(* Logix 5000 project; controller PLC_MCC1201_220AP1 vendor 1 type 14 code 164 rev 35.11; software revision 35.00; part 19 of 25 *)
(* tags used below, declared in another part *)
   TMP_xSimulationMode : BOOL;
   AFI : ALIAS FOR B3[7].15;
   AMAX_LEHR_SPD : ALIAS FOR I[81];
   C5 : COUNTER[100];
   C5_ACTIVE_LAMP : ALIAS FOR N54[264].0;
   C5_NTH_IN_LMP : ALIAS FOR N54[264].10;
   C5_NTH_IN_PE : ALIAS FOR N54[264].6;
   C5_NTH_OUT_LMP : ALIAS FOR N54[264].9;
   C5_NTH_OUT_PE : ALIAS FOR N54[264].5;
   C5_STH_IN_LMP : ALIAS FOR N54[264].12;
   C5_STH_IN_PE : ALIAS FOR N54[264].8;
   C5_STH_OUT_LMP : ALIAS FOR N54[264].11;
   C5_STH_OUT_PE : ALIAS FOR N54[264].7;
   CR1_DNET_SS1 : ALIAS FOR N179[18];
   CR1_DNET_SS2 : ALIAS FOR N179[30];
   DRIVE_FAULT_PRESENT : BOOL;
   F96 : REAL[50];
   HMI_Alarm_Presence : BOOL;   // HMI_Alarm_Presence
   HMI_Alarms_0 : BOOL[32];   // HMI Alarms
   HMI_Alarms_1 : BOOL[32];   // HMI Alarms
   HMI_Alarms_2 : BOOL[32];   // HMI Alarms
   HMI_Alarms_3 : BOOL[32];   // HMI Alarms
   HMI_Alarms_4 : BOOL[32];   // HMI Alarms
   HMI_Alarms_5 : BOOL[32];   // HMI Alarms
   HMI_Alarms_6 : BOOL[32];   // HMI Alarms
   HMI_Alarms_7 : BOOL[32];   // HMI Alarms
   HMI_Alarms_8 : BOOL[32];   // HMI Alarms
   HMI_Alarms_9 : BOOL[32];   // HMI Alarms
   HMI_MAN_CMD_WR : UDT_MAN_CMD_WR;
   I : INT[128];
   LEHRSPD_CURRENT : ALIAS FOR N98[5];
   M203DROP : MAC_DROPCONV;
   M205BREAKER : MAC_BREAKER;
   M225 : MAC_EMERGENCYXCUT;
   N11 : DINT[1000];
   N11_HOST : INT[1000];
   N12 : DINT[1000];
   N12_HOST : INT[1000];
   N14 : DINT[1000];
   N14_HOST : INT[1000];
   N179 : DINT[600];
   N500 : DINT[24];
   N501 : DINT[25];
   N502 : DINT[25];
   N504 : DINT[25];
   N505 : DINT[25];
   N507 : DINT[25];
   N53 : DINT[10];
   N53_HOST : INT[10];
   N54 : DINT[501];
   N54_HOST : INT[501];
   O : INT[128];
   ProducedToCullet : UDT_PRODUCED_CULLET;
   ProducedToMCC1300 : UDT_PRODUCED_NEXT;
   R509 : CONTROL[2];
   R509_000_POS : ALIAS FOR R509[0].POS;
   R509_001_POS : ALIAS FOR R509[1].POS;
   S : INT[128];
   Sbr_IN_dDataLength : DINT;
   Status : INT;   // INT tag to retrieve Status value through GSV created during conversion
   T160 : TIMER[100];
   TMP_dIndex : DINT;
   TMP_Index : DINT;
   TMP_xAlwaysOFF : BOOL;
   To_Cullet : DINT[10];
   W_APC_ACTIVE : ALIAS FOR W_B3[0].10;
   W_B3 : DINT[7];
   W_C5 : COUNTER[1];
   W_CB1_AUXILLARY : ALIAS FOR W_I[8].12;
   W_CB1_START : ALIAS FOR W_O[10].1;
   W_CB2_AUXILLARY : ALIAS FOR W_I[8].11;
   W_CB2_START : ALIAS FOR W_O[10].3;
   W_CONV_MSG_N7_0 : MESSAGE;   // IFE1_BTW_CNT
   W_CONV_MSG_N7_120 : MESSAGE;   // OFE1_CONTROL
   W_CONV_MSG_N7_160 : MESSAGE;   // OFE1_BTR_CONTRO
   W_CONV_MSG_N7_200 : MESSAGE;   // OFE2_CONTROL
   W_CONV_MSG_N7_240 : MESSAGE;   // OFE2_BTR_CONTRO
   W_CONV_MSG_N7_280 : MESSAGE;   // OFE3_CONTROL
   W_CONV_MSG_N7_32 : MESSAGE;   // IFE1_BTR
   W_CONV_MSG_N7_320 : MESSAGE;   // OFE3_BTR_CONTRL
   W_CONV_MSG_N7_360 : MESSAGE;   // OFE4_CONTROL
   W_CONV_MSG_N7_400 : MESSAGE;   // OFE4_BTR_CONTRL
   W_CONV_MSG_N7_60 : MESSAGE;   // IFE2_CONTROL
   W_CONV_MSG_N7_92 : MESSAGE;   // IFE2_BTR
   W_CONV_PID_N7_440 : PID;   // Receiving Tank Level Control
   W_CONV_PID_N7_470 : PID;   // Washer Water Pressure Cntrl Valve Position
   W_CONV_PID_N7_500 : PID;   // Dryer Room Airflow (CB2) Fan Actuator Control
   W_CONV_PID_N7_530 : PID;   // Blower CB1 Static Pressure Fan Actuator Control
   W_CONV_PID_N7_560 : PID;   // RO Heating Coil Temp. Control (HC1)
   W_CONV_PID_N7_590 : PID;   // Eclipse Heating Coil Temp. Control
   W_CP1_ENABLE : ALIAS FOR W_B3[0].5;
   W_CP1A_START : ALIAS FOR W_O[10].5;
   W_CP1A_STATUS : ALIAS FOR W_I[8].7;
   W_CP1B_START : ALIAS FOR W_O[10].7;
   W_CP1B_STATUS : ALIAS FOR W_I[8].6;
   W_CP2A_START : ALIAS FOR W_O[10].9;
   W_CP2A_STAT : ALIAS FOR W_I[8].4;
   W_CP2B_START : ALIAS FOR W_O[10].11;
   W_CP2B_STAT : ALIAS FOR W_I[8].3;
   W_DRV_OUTPUT : ALIAS FOR W_N7[380];
   W_DRYER_AIR_FLOW : ALIAS FOR W_N7[108];
   W_EMER_STOP : ALIAS FOR W_I[8].13;
   W_EMER_STOP_LIGHT : ALIAS FOR W_O[10].10;
   W_FLOW_ENABLE : ALIAS FOR W_B3[0].9;
   W_HEATING_AIR_ST : ALIAS FOR W_N7[107];
   W_I : INT[32];
   W_INT_FOR_BCD1 : ALIAS FOR W_N7[911];
   W_LEVEL_SENSOR : ALIAS FOR W_N7[109];
   W_LL_CP1 : ALIAS FOR W_I[8].14;
   W_LL_CP2 : ALIAS FOR W_I[8].15;
   W_LOG_SHUTDOWN : ALIAS FOR W_I[8].0;
   W_N7 : DINT[933];
   W_O : INT[32];
   W_OUT_FROM_PID : ALIAS FOR W_N7[907];
   W_PID_BCD_TCD2 : ALIAS FOR W_N7[913];
   W_PID_TO_OUTPUT : ALIAS FOR W_N7[903];
   W_PS1_SWITCH : ALIAS FOR W_I[8].8;
   W_PWT_HIGH_LIMIT : ALIAS FOR W_I[8].2;
   W_RECIEVING_LEVEL : ALIAS FOR W_I[8].9;
   W_RO_SIG_START : ALIAS FOR W_B3[6].4;
   W_RO_START : ALIAS FOR W_O[10].13;
   W_RUN_WASHER : ALIAS FOR W_B3[0].2;
   W_SHUTDOWN_LATCH : ALIAS FOR W_B3[0].1;
   W_SIG_CP1A_START : ALIAS FOR W_B3[0].6;
   W_SIG_CP1B_START : ALIAS FOR W_B3[0].7;
   W_SIG_CP2A_START : ALIAS FOR W_B3[0].3;
   W_SIG_CP2B_START : ALIAS FOR W_B3[0].4;
   W_T4 : TIMER[101];
   W_TCD1_OUTPUT : ALIAS FOR W_N7[222];
   W_TCD2_OUTPUT : ALIAS FOR W_N7[223];
   W_TT8_INPUT : ALIAS FOR W_N7[912];
   W_TT8_RAW_DATA : ALIAS FOR W_N7[53];
   W_WARNING_LIGHT : ALIAS FOR W_O[10].8;
   Z200 : MAC_Zone_ML;
(* MainProgram, continued *)

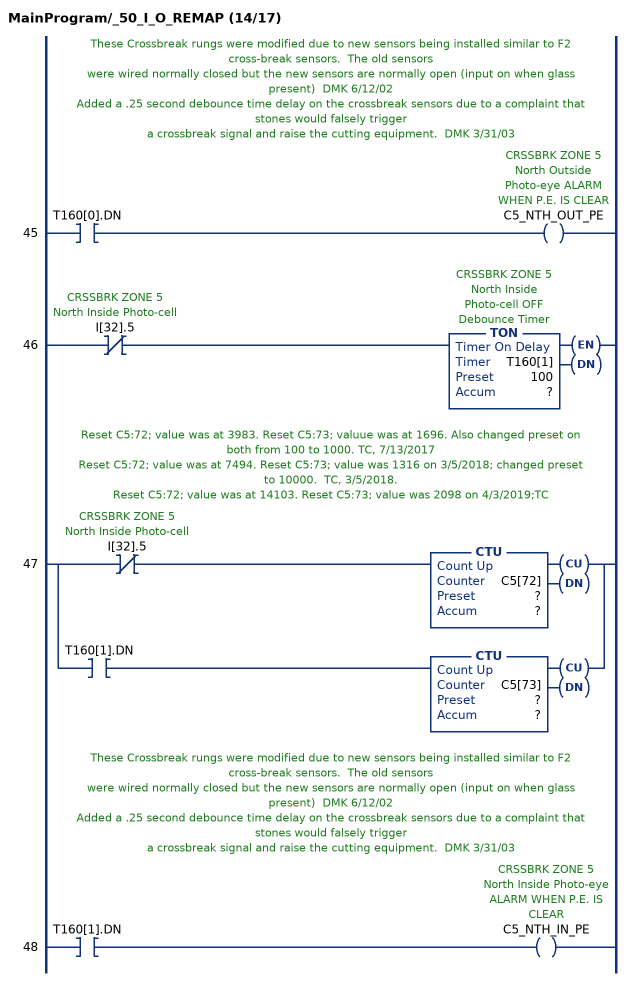
   [picture p306: MainProgram/_50_I_O_REMAP rungs 45-48]
   // These Crossbreak rungs were modified due to new sensors being installed similar to F2 cross-break sensors.  The old sensors
   // were wired normally closed but the new sensors are normally open (input on when glass present)  DMK 6/12/02
   // Added a .25 second debounce time delay on the crossbreak sensors due to a complaint that stones would falsely trigger
   // a crossbreak signal and raise the cutting equipment.  DMK 3/31/03
   45: XIC(T160[0].DN)OTE(C5_NTH_OUT_PE);
   46: XIO(I[32].5)TON(T160[1],?,?);
   // Reset C5:72; value was at 3983. Reset C5:73; valuue was at 1696. Also changed preset on both from 100 to 1000. TC, 7/13/2017
   //                                                                                                                                                       Reset C5:72; value was at 7494. Reset C5:73; value was 1316 on 3/5/2018; changed preset to 10000.  TC, 3/5/2018.
   //                                                                                                                                                                      Reset C5:72; value was at 14103. Reset C5:73; value was 2098 on 4/3/2019;TC
   47: [XIO(I[32].5) CTU(C5[72],?,?) ,XIC(T160[1].DN) CTU(C5[73],?,?) ];
   // These Crossbreak rungs were modified due to new sensors being installed similar to F2 cross-break sensors.  The old sensors
   // were wired normally closed but the new sensors are normally open (input on when glass present)  DMK 6/12/02
   // Added a .25 second debounce time delay on the crossbreak sensors due to a complaint that stones would falsely trigger
   // a crossbreak signal and raise the cutting equipment.  DMK 3/31/03
   48: XIC(T160[1].DN)OTE(C5_NTH_IN_PE);
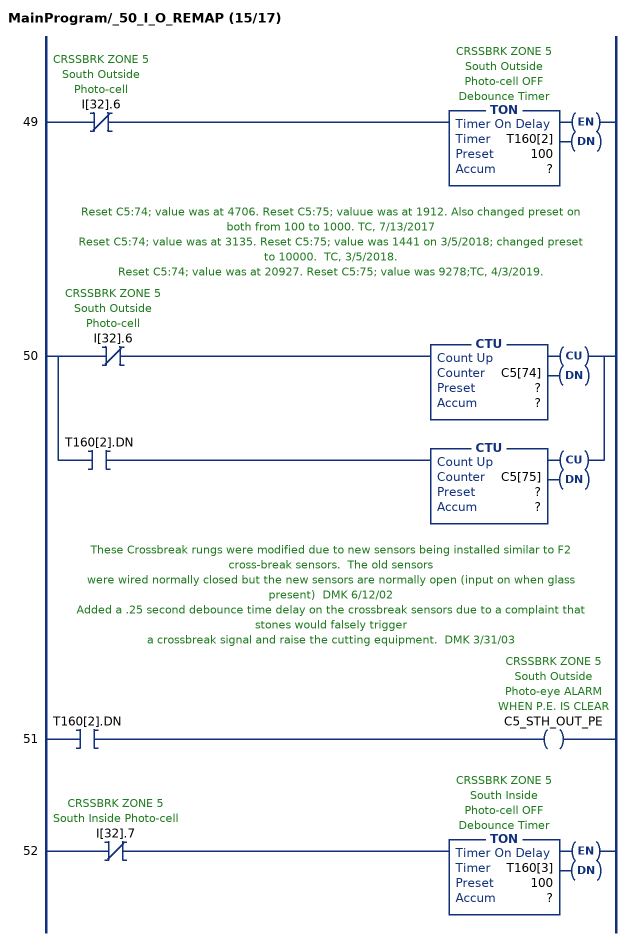
   49: XIO(I[32].6)TON(T160[2],?,?);
   // Reset C5:74; value was at 4706. Reset C5:75; valuue was at 1912. Also changed preset on both from 100 to 1000. TC, 7/13/2017
   //                                                                                                                                                                  Reset C5:74; value was at 3135. Reset C5:75; value was 1441 on 3/5/2018; changed preset to 10000.  TC, 3/5/2018.
   //                                                                                                                                                                                          Reset C5:74; value was at 20927. Reset C5:75; value was 9278;TC, 4/3/2019.
   50: [XIO(I[32].6) CTU(C5[74],?,?) ,XIC(T160[2].DN) CTU(C5[75],?,?) ];
   // These Crossbreak rungs were modified due to new sensors being installed similar to F2 cross-break sensors.  The old sensors
   // were wired normally closed but the new sensors are normally open (input on when glass present)  DMK 6/12/02
   // Added a .25 second debounce time delay on the crossbreak sensors due to a complaint that stones would falsely trigger
   // a crossbreak signal and raise the cutting equipment.  DMK 3/31/03
   51: XIC(T160[2].DN)OTE(C5_STH_OUT_PE);
   52: XIO(I[32].7)TON(T160[3],?,?);
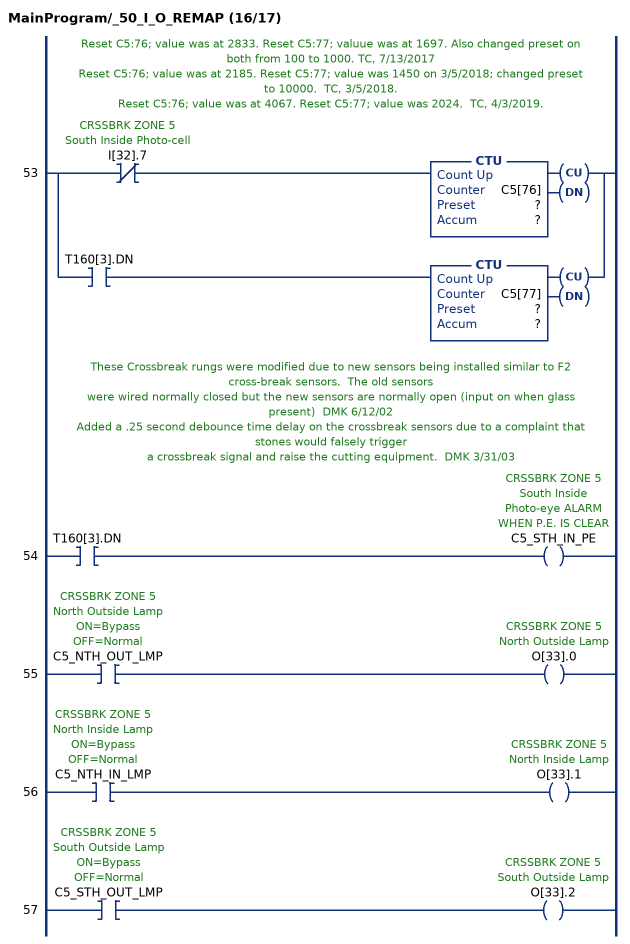
   // Reset C5:76; value was at 2833. Reset C5:77; valuue was at 1697. Also changed preset on both from 100 to 1000. TC, 7/13/2017
   //                                                                                                                                                     Reset C5:76; value was at 2185. Reset C5:77; value was 1450 on 3/5/2018; changed preset to 10000.  TC, 3/5/2018.
   //                                                                                                                                                                               Reset C5:76; value was at 4067. Reset C5:77; value was 2024.  TC, 4/3/2019.
   53: [XIO(I[32].7) CTU(C5[76],?,?) ,XIC(T160[3].DN) CTU(C5[77],?,?) ];
   // These Crossbreak rungs were modified due to new sensors being installed similar to F2 cross-break sensors.  The old sensors
   // were wired normally closed but the new sensors are normally open (input on when glass present)  DMK 6/12/02
   // Added a .25 second debounce time delay on the crossbreak sensors due to a complaint that stones would falsely trigger
   // a crossbreak signal and raise the cutting equipment.  DMK 3/31/03
   54: XIC(T160[3].DN)OTE(C5_STH_IN_PE);
   55: XIC(C5_NTH_OUT_LMP)OTE(O[33].0);
   56: XIC(C5_NTH_IN_LMP)OTE(O[33].1);
   57: XIC(C5_STH_OUT_LMP)OTE(O[33].2);
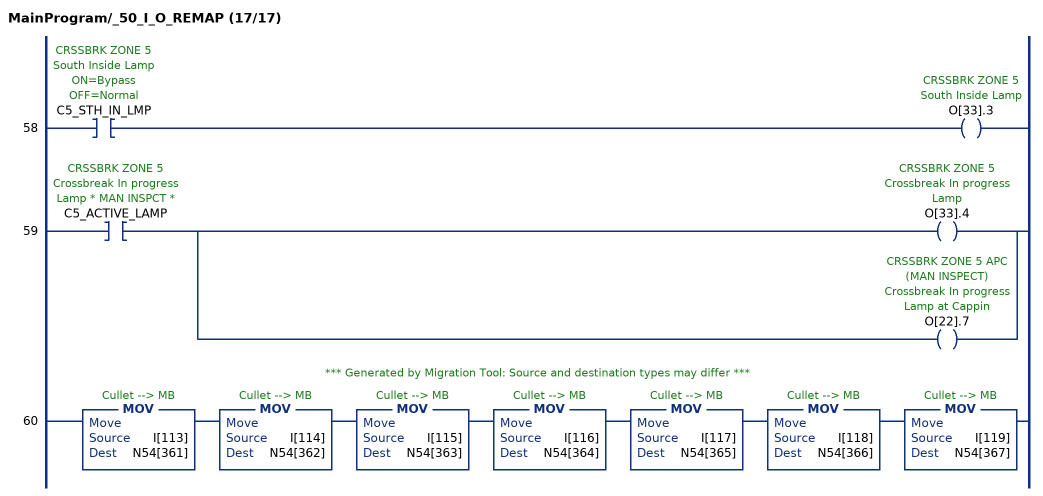
   58: XIC(C5_STH_IN_LMP)OTE(O[33].3);
   59: XIC(C5_ACTIVE_LAMP)[OTE(O[33].4) ,OTE(O[22].7) ];
   // *** Generated by Migration Tool: Source and destination types may differ ***
   60: MOV(I[113],N54[361])MOV(I[114],N54[362])MOV(I[115],N54[363])MOV(I[116],N54[364])MOV(I[117],N54[365])MOV(I[118],N54[366])MOV(I[119],N54[367]);
END_ROUTINE

ROUTINE _51_LADDER   (* ladder *)
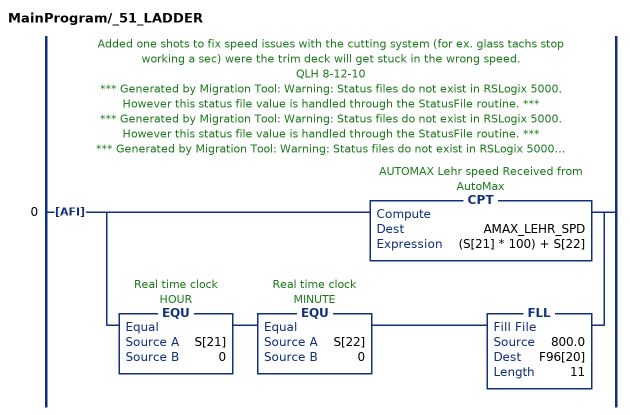
   // Added one shots to fix speed issues with the cutting system (for ex. glass tachs stop working a sec) were the trim deck will get stuck in the wrong speed.
   // QLH 8-12-10
   // *** Generated by Migration Tool: Warning: Status files do not exist in RSLogix 5000. However this status file value is handled through the StatusFile routine. ***
   // *** Generated by Migration Tool: Warning: Status files do not exist in RSLogix 5000. However this status file value is handled through the StatusFile routine. ***
   // *** Generated by Migration Tool: Warning: Status files do not exist in RSLogix 5000. However this status file value is handled through the StatusFile routine. ***
   // *** Generated by Migration Tool: Warning: Status files do not exist in RSLogix 5000. However this status file value is handled through the StatusFile routine. ***
   0: AFI()[CPT(AMAX_LEHR_SPD,(S[21] * 100) + S[22]) ,EQU(S[21],0) EQU(S[22],0) FLL(800.0,F96[20],11) ];
END_ROUTINE

ROUTINE _811_HOST_MOVE   (* structured text *)
   
   //Input
   SBR(Sbr_IN_dDataLength);
   
   FOR TMP_dIndex := 0 TO Sbr_IN_dDataLength - 1 DO
   	N11_HOST[TMP_dIndex] := N11[TMP_dIndex];
   END_FOR;
   
END_ROUTINE

ROUTINE _812_HOST_MOVE   (* structured text *)
   
   //Input
   SBR(Sbr_IN_dDataLength);
   
   FOR TMP_dIndex := 0 TO Sbr_IN_dDataLength - 1 DO
   	N12[TMP_dIndex] := N12_HOST[TMP_dIndex];
   END_FOR;
   
END_ROUTINE

ROUTINE _814_HOST_MOVE   (* structured text *)
   
   
   //Input
   SBR(Sbr_IN_dDataLength);
   
   FOR TMP_dIndex := 0 TO Sbr_IN_dDataLength - 1 DO
   	N14[TMP_dIndex] := N14_HOST[TMP_dIndex];
   END_FOR;
   
END_ROUTINE

ROUTINE _853_HOST_MOVE   (* structured text *)
   
   //Input
   SBR(Sbr_IN_dDataLength);
   
   FOR TMP_dIndex := 0 TO Sbr_IN_dDataLength - 1 DO
   	N53[TMP_dIndex] := N53_HOST[TMP_dIndex];
   END_FOR;
   
END_ROUTINE

ROUTINE _854_HOST_MOVE   (* structured text *)
   
   //Input
   SBR(Sbr_IN_dDataLength);
   
   FOR TMP_dIndex := 0 TO Sbr_IN_dDataLength - 1 DO
   	N54_HOST[TMP_dIndex] := N54[TMP_dIndex];
   END_FOR;
   
END_ROUTINE

ROUTINE _880_HMI_Mapping   (* structured text *)
   
   // Alarm maps for HMI
   TMP_Index:= 0;
   FOR TMP_Index := 0 TO 15 DO
   	//HMI_Alarms_0[TMP_Index]:= N11[62].[TMP_Index];
   	//HMI_Alarms_1[TMP_Index]:= N11[64].[TMP_Index];
   	HMI_Alarms_0[TMP_Index]:= 0;
   	HMI_Alarms_1[TMP_Index]:= 0;
   	HMI_Alarms_2[TMP_Index]:= 0;
   	HMI_Alarms_3[TMP_Index]:= 0;
   	HMI_Alarms_4[TMP_Index]:= 0;
   	HMI_Alarms_5[TMP_Index]:= 0;
   	HMI_Alarms_6[TMP_Index]:= 0;
   	HMI_Alarms_7[TMP_Index]:= 0;
   	HMI_Alarms_8[TMP_Index]:= 0;
   	HMI_Alarms_9[TMP_Index]:= 0;
   	//HMI_Alarms_2[TMP_Index]:= NOT N11[22].[TMP_Index];
   	//HMI_Alarms_3[TMP_Index]:= NOT N11[23].[TMP_Index];
   END_FOR;
   FOR TMP_Index := 16 TO 31 DO
   	HMI_Alarms_0[TMP_Index]:= 0;
   	HMI_Alarms_1[TMP_Index]:= 0;
   	HMI_Alarms_2[TMP_Index]:= 0;
   	HMI_Alarms_3[TMP_Index]:= 0;
   	HMI_Alarms_4[TMP_Index]:= 0;
   	HMI_Alarms_5[TMP_Index]:= 0;
   	HMI_Alarms_6[TMP_Index]:= 0;
   	HMI_Alarms_7[TMP_Index]:= 0;
   	HMI_Alarms_8[TMP_Index]:= 0;
   	HMI_Alarms_9[TMP_Index]:= 0;
   END_FOR;
   
   (*
   HMI_Alarms_0[0] := NOT N11[20].0;
   HMI_Alarms_0[1] := NOT N11[20].1;
   HMI_Alarms_0[2] := NOT N11[20].2;
   HMI_Alarms_0[3] := NOT N11[20].3;
   HMI_Alarms_0[4] := 0;
   HMI_Alarms_0[5] := NOT N11[20].5;
   HMI_Alarms_0[6] := NOT N11[20].6;
   HMI_Alarms_0[7] := NOT N11[20].7;
   HMI_Alarms_0[8] := N11[20].8;
   HMI_Alarms_0[9] := N11[20].9;
   HMI_Alarms_0[10] := NOT N11[20].10;
   HMI_Alarms_0[11] := NOT N11[20].11;
   HMI_Alarms_0[12] := NOT N11[20].12;
   HMI_Alarms_0[13] := NOT N11[20].13;
   HMI_Alarms_0[14] := N11[20].14;
   HMI_Alarms_0[15] := 0;
   
   HMI_Alarms_2[0] := NOT N11[22].0;
   HMI_Alarms_2[1] := NOT N11[22].1;
   HMI_Alarms_2[2] := NOT N11[22].2;
   HMI_Alarms_2[3] := NOT N11[22].3;
   HMI_Alarms_2[4] := NOT N11[22].4;
   HMI_Alarms_2[5] := NOT N11[22].5;
   HMI_Alarms_2[6] := NOT N11[22].6;
   HMI_Alarms_2[7] := NOT N11[22].7;
   HMI_Alarms_2[8] := NOT N11[22].8;
   HMI_Alarms_2[9] := NOT N11[22].9;
   HMI_Alarms_2[10] := NOT N11[22].10;
   HMI_Alarms_2[11] := NOT N11[22].11;
   HMI_Alarms_2[12] := NOT N11[22].12;
   HMI_Alarms_2[13] := NOT N11[22].13;
   HMI_Alarms_2[14] := 0;
   HMI_Alarms_2[15] := 0;
   
   HMI_Alarms_3[0] := NOT N11[23].0;
   HMI_Alarms_3[1] := NOT N11[23].1;
   HMI_Alarms_3[2] := NOT N11[23].2;
   HMI_Alarms_3[3] := NOT N11[23].3;
   HMI_Alarms_3[4] := NOT N11[23].4;
   HMI_Alarms_3[5] := NOT N11[23].5;
   HMI_Alarms_3[6] := NOT N11[23].6;
   HMI_Alarms_3[7] := NOT N11[23].7;
   HMI_Alarms_3[8] := NOT N11[23].8;
   HMI_Alarms_3[9] := NOT N11[23].9;
   HMI_Alarms_3[10] := NOT N11[23].10;
   HMI_Alarms_3[11] := NOT N11[23].11;
   HMI_Alarms_3[12] := NOT N11[23].12;
   HMI_Alarms_3[13] := NOT N11[23].13;
   HMI_Alarms_3[14] := 0;
   HMI_Alarms_3[15] := 0;
   
   HMI_Alarms_9[0] := M316M1_IN.Faulted;
   HMI_Alarms_9[1] := M317M1_IN.Faulted;
   HMI_Alarms_9[2] := M317M2_IN.Faulted;
   HMI_Alarms_9[3] := M317M3_IN.Faulted;
   HMI_Alarms_9[4] := M317M4_IN.Faulted;
   HMI_Alarms_9[5] := M317M5_IN.Faulted;
   HMI_Alarms_9[6] := M317M6_IN.Faulted;
   HMI_Alarms_9[7] := M318M1_IN.Faulted;
   HMI_Alarms_9[8] := M318AM1_IN.Faulted;
   HMI_Alarms_9[9] := M318BM1_IN.Faulted;
   HMI_Alarms_9[10] := M318BM2_IN.Faulted;
   HMI_Alarms_9[11] := M318BM3_IN.Faulted;
   HMI_Alarms_9[12] := M318BM4_IN.Faulted;
   HMI_Alarms_9[13] := M391M1_IN.Faulted;
   *)
   
   // Alarm presence for HMI
   HMI_Alarm_Presence := 0;
   TMP_Index:= 0;
   FOR TMP_Index := 0 TO 31 DO
   	IF HMI_Alarms_0[TMP_Index] OR HMI_Alarms_1[TMP_Index] OR HMI_Alarms_2[TMP_Index] OR HMI_Alarms_3[TMP_Index] OR HMI_Alarms_4[TMP_Index] OR HMI_Alarms_5[TMP_Index] THEN
   		HMI_Alarm_Presence := 1;
   	END_IF;
   	IF HMI_Alarms_6[TMP_Index] OR HMI_Alarms_7[TMP_Index] OR HMI_Alarms_8[TMP_Index] OR HMI_Alarms_9[TMP_Index] THEN
   		HMI_Alarm_Presence := 1;
   	END_IF;
   END_FOR;
   
   //// Logic to make horn sound for drives fault
   //DRIVE_FAULT_PRESENT := 0;
   //FOR TMP_Index := 0 TO 8 BY 1 DO
   //	IF N11[62].[TMP_Index] THEN
   //		DRIVE_FAULT_PRESENT := 1;
   //	END_IF;
   //END_FOR;
   
   (*
   // Photocell maps for HMI
   HMI_ProxySwitch[0] := I[2].0;
   HMI_ProxySwitch[1] := I[2].1;
   HMI_ProxySwitch[2] := I[2].2;
   HMI_ProxySwitch[3] := I[2].3;
   HMI_ProxySwitch[4] := I[2].4;
   HMI_ProxySwitch[5] := I[2].5;
   HMI_ProxySwitch[6] := I[2].6;
   HMI_ProxySwitch[7] := I[2].7;
   HMI_ProxySwitch[8] := I[2].8;
   HMI_ProxySwitch[9] := I[2].9;
   HMI_ProxySwitch[10] := I[2].10;
   HMI_ProxySwitch[11] := I[2].11;
   HMI_ProxySwitch[12] := I[2].12;
   HMI_ProxySwitch[13] := I[2].13;
   HMI_ProxySwitch[14] := I[2].14;
   HMI_ProxySwitch[15] := I[2].15;
   
   // Photocell maps for HMI
   HMI_Photocells[0] := I[3].0;
   HMI_Photocells[1] := I[3].1;
   HMI_Photocells[2] := I[3].2;
   HMI_Photocells[3] := I[3].3;
   HMI_Photocells[4] := I[3].4;
   HMI_Photocells[5] := I[3].5;
   HMI_Photocells[6] := I[3].6;
   HMI_Photocells[7] := I[3].7;
   HMI_Photocells[8] := I[3].8;
   HMI_Photocells[9] := I[3].9;
   HMI_Photocells[10] := I[3].10;
   HMI_Photocells[11] := I[3].11;
   HMI_Photocells[12] := I[3].12;
   HMI_Photocells[13] := I[3].13;
   HMI_Photocells[14] := I[3].14;
   HMI_Photocells[15] := I[3].15;
   
   HMI_Photocells[16] := I[5].8;
   HMI_Photocells[17] := I[5].9;
   
   //All commands
   I[21].15 := HMI_MAN_CMD_WR.CONV_Manual_ALL;
   I[23].15 := HMI_MAN_CMD_WR.CONV_Man_ALL_FWD;
   I[25].15 := HMI_MAN_CMD_WR.CONV_Man_ALL_REV;
   
   //M316M1 Roll Conveyor M4CM01
   I[20].0 := HMI_MAN_CMD_WR.M316M1_Manual;
   I[22].0 := HMI_MAN_CMD_WR.M316M1_ManFWD;
   I[24].0 := HMI_MAN_CMD_WR.M316M1_ManREV;
   
   //M317M1 Roll Conveyor Zone 1 M4CM02
   I[20].1 := HMI_MAN_CMD_WR.M317M1_Manual;
   I[22].1 := HMI_MAN_CMD_WR.M317M1_ManFWD;
   I[24].1 := HMI_MAN_CMD_WR.M317M1_ManREV;
   
   //M317M2 Lifting Zone 1 M4CM03
   I[20].2 := HMI_MAN_CMD_WR.M317M2_Manual;
   I[22].2 := HMI_MAN_CMD_WR.M317M2_ManFWD;
   I[24].2 := HMI_MAN_CMD_WR.M317M2_ManREV;
   
   //M317M3 Lifting Zone 2 M4CM04
   I[20].3 := HMI_MAN_CMD_WR.M317M3_Manual;
   I[22].3 := HMI_MAN_CMD_WR.M317M3_ManFWD;
   I[24].3 := HMI_MAN_CMD_WR.M317M3_ManREV;
   
   //M317M4 Roll Conveyor Zone 2 M4CM05
   I[20].4 := HMI_MAN_CMD_WR.M317M4_Manual;
   I[22].4 := HMI_MAN_CMD_WR.M317M4_ManFWD;
   I[24].4 := HMI_MAN_CMD_WR.M317M4_ManREV;
   
   //M317M5 Wheel Conveyor Zone 1 M4CM06
   I[20].5 := HMI_MAN_CMD_WR.M317M5_Manual;
   I[22].5 := HMI_MAN_CMD_WR.M317M5_ManFWD;
   I[24].5 := HMI_MAN_CMD_WR.M317M5_ManREV;
   
   //M317M6 Wheel Conveyor Zone 2 M4CM07
   I[20].6 := HMI_MAN_CMD_WR.M317M6_Manual;
   I[22].6 := HMI_MAN_CMD_WR.M317M6_ManFWD;
   I[24].6 := HMI_MAN_CMD_WR.M317M6_ManREV;
   
   //M318M1 Roll Conveyor M4CM08
   I[20].7 := HMI_MAN_CMD_WR.M318M1_Manual;
   I[22].7 := HMI_MAN_CMD_WR.M318M1_ManFWD;
   I[24].7 := HMI_MAN_CMD_WR.M318M1_ManREV;
   
   //M318AM1 Roll Conveyor M4CM09
   I[20].8 := HMI_MAN_CMD_WR.M318AM1_Manual;
   I[22].8 := HMI_MAN_CMD_WR.M318AM1_ManFWD;
   I[24].8 := HMI_MAN_CMD_WR.M318AM1_ManREV;
   
   //M318BM1 Roll Conveyor Zone 1 M4CM10
   I[20].9 := HMI_MAN_CMD_WR.M318BM1_Manual;
   I[22].9 := HMI_MAN_CMD_WR.M318BM1_ManFWD;
   I[24].9 := HMI_MAN_CMD_WR.M318BM1_ManREV;
   
   //M318BM2 Lifting Zone 1 M4CM11
   I[20].10 := HMI_MAN_CMD_WR.M318BM2_Manual;
   I[22].10 := HMI_MAN_CMD_WR.M318BM2_ManFWD;
   I[24].10 := HMI_MAN_CMD_WR.M318BM2_ManREV;
   
   //M318BM3 Lifting Zone 2 M4CM12
   I[20].11 := HMI_MAN_CMD_WR.M318BM3_Manual;
   I[22].11 := HMI_MAN_CMD_WR.M318BM3_ManFWD;
   I[24].11 := HMI_MAN_CMD_WR.M318BM3_ManREV;
   
   //M318BM4 Roll Conveyor Zone 2 M4CM13
   I[20].12 := HMI_MAN_CMD_WR.M318BM4_Manual;
   I[22].12 := HMI_MAN_CMD_WR.M318BM4_ManFWD;
   I[24].12 := HMI_MAN_CMD_WR.M318BM4_ManREV;
   
   //M391M1 Wheel Conveyor (Sample Table) M4CM14
   I[20].13 := HMI_MAN_CMD_WR.M391M1_Manual;
   I[22].13 := HMI_MAN_CMD_WR.M391M1_ManFWD;
   I[24].13 := HMI_MAN_CMD_WR.M391M1_ManREV;
   I[22].14 := HMI_MAN_CMD_WR.M391_ManRAISE;
   I[24].14 := HMI_MAN_CMD_WR.M391_ManLOWER;
   *)
   
END_ROUTINE

ROUTINE _990_Output_Mapping   (* structured text *)
   
   //OUTPUT
   
   //MCC1201
   A152AP1:14:O.Pt00.Data := Z200.OUTPUT_xMainEmergencyLamp;
   A152AP1:14:O.Pt01.Data := Z200.OUTPUT_xUPSEmergencyLamp;
   A152AP1:14:O.Pt02.Data := Z200.OUTPUT_xMCCSafetyLamp;
   
   //Alarms signalling
   A152AP1:15:O.Pt03.Data := Z200.OUTPUT_xUPSEmergencyLamp;
   A152AP1:15:O.Pt06.Data := Z200.OUTPUT_xAcousticAlarm;
   A152AP1:15:O.Pt07.Data := Z200.OUTPUT_xUPSEmergencyLamp;
   A152AP1:15:O.Pt11.Data := Z200.OUTPUT_xMainEmergencyLamp;
   A152AP1:15:O.Pt12.Data := Z200.OUTPUT_xMainEmergencyLamp;
   A152AP1:16:O.Pt01.Data := Z200.OUTPUT_xUPSEmergencyLamp;
   A152AP1:16:O.Pt11.Data := Z200.OUTPUT_xUPSEmergencyLamp;
   
   //M203DROP
   A152AP1:15:O.Pt00.Data := M203DROP.OUTPUT_xRollerLifting;
   A152AP1:15:O.Pt01.Data := M203DROP.OUTPUT_xDescentDrop;
   A152AP1:15:O.Pt02.Data := M203DROP.OUTPUT_xRiseDrop;
   A152AP1:15:O.Pt04.Data := M203DROP.OUTPUT_xHLDoorOpenOpSide;
   A152AP1:15:O.Pt05.Data := M203DROP.OUTPUT_xHLUpDownPushbutton;
   A152AP1:15:O.Pt08.Data := M203DROP.OUTPUT_xHLDoorOpenFarSide;
   A152AP1:15:O.Pt09.Data := M203DROP.OUTPUT_xHLUpDownPushbutton;
   
   //M225 EMERGENCY XCUT
   A152AP1:16:O.Pt00.Data := M225.OUTPUT_xUnlockDoorOpSide;
   A152AP1:16:O.Pt02.Data := M225.OUTPUT_xAreaAccessRequestFarSide;
   A152AP1:16:O.Pt05.Data := M225.OUTPUT_xUnlockDoorFarSide;
   A152AP1:16:O.Pt06.Data := M225.OUTPUT_xMachineReady;
   A152AP1:16:O.Pt07.Data := M225.OUTPUT_xMachineToMaintenance;
   A152AP1:16:O.Pt08.Data := M225.OUTPUT_xMachineOutOfOrder;
   A152AP1:18:O.Pt00.Data := M225.OUTPUT_xCuttingHeadDescent;
   A152AP1:18:O.Pt01.Data := M225.OUTPUT_xLubrication;
   A152AP1:18:O.Pt02.Data := M225.OUTPUT_xAirActivation;
   
   //CS4225 EMERGENCY XCUT CONSOLLE
   A152AP1:16:O.Pt12.Data := M225.OUTPUT_xAreaAccessRequestOpSide;
   A152AP1:16:O.Pt13.Data := M225.OUTPUT_xAutomatic;
   A152AP1:16:O.Pt14.Data := M225.OUTPUT_xStartCut;
   A152AP1:16:O.Pt15.Data := M225.OUTPUT_xStopCut;
   
   //M205BREAKER
   A152AP1:13:O.Pt00.Data := M205BREAKER.OUTPUT_xBreakerRun;
   
   //M225
   A152AP1:13:O.Pt01.Data := M225.OUTPUT_xCarriageOverstroke;
   
   
   // MAPPING PREVIOUS PROGRAM OUTPUTS
   
   //HORN / CHILLED WATER / APC / SUBSURFACE / ISRA 5D
   A152AP1:14:O.Pt03.Data := I[20].3; //PLC ALARM HORN RELAY
   A152AP1:14:O.Pt04.Data := I[20].4; //North Chilled Water Blower Start VFD
   A152AP1:14:O.Pt05.Data := I[20].5; //North Chilled Water Blower Start LT I02104 PB
   A152AP1:14:O.Pt06.Data := I[20].6; //North Chilled Water VFD Stop
   A152AP1:14:O.Pt07.Data := I[20].0; //South Chilled Water Blower Start VFD
   A152AP1:14:O.Pt08.Data := I[20].1; //South Chilled Water Blower Start LT I02112 PB
   A152AP1:14:O.Pt09.Data := I[20].2; //South Chilled Water VFD Stop
   A152AP1:14:O.Pt10.Data := I[20].8; //LUCOR MACHINE OPERATE (APC CONTACTORS?)
   A152AP1:14:O.Pt11.Data := I[20].11; //SUB-SURFACE Cutters Raise for Crossbreak Relay
   A152AP1:14:O.Pt12.Data := I[20].12; //ISRA 5D System Cut Signal
   A152AP1:14:O.Pt13.Data := I[20].13; //ISRA 5D System QC Request Signal
   
   // CROSSBREAK ZONE 1
   CB_1CS:1:O.0 := O[25].0; //CRSSBRK ZONE 1 North Outside Lamp
   CB_1CS:1:O.1 := O[25].1; //CRSSBRK ZONE 1 North Inside Lamp
   CB_1CS:1:O.2 := O[25].2; //CRSSBRK ZONE 1 South Outside Lamp
   CB_1CS:1:O.3 := O[25].3; //CRSSBRK ZONE 1 South Inside Lamp
   CB_1CS:1:O.4 := O[25].4; //CRSSBRK ZONE 1 Crossbreak In progress Lamp
   CB_1CS:1:O.5 := O[25].5; //M37B Conv Forward Pilot Light
   CB_1CS:1:O.6 := O[25].6; //M37B Conv Reverse Pilot Light
   CB_1CS:1:O.7 := O[25].7; //M47B Conv Forward Pilot Light
   CB_1CS:1:O.8 := O[25].8; //M47B Conv Reverse Pilot Light
   CB_1CS:1:O.9 := O[25].9; //spare
   CB_1CS:1:O.10 := O[25].10; //spare
   CB_1CS:1:O.11 := O[25].11; //spare
   CB_1CS:1:O.12 := O[25].12; //spare
   CB_1CS:1:O.13 := O[25].13; //spare
   CB_1CS:1:O.14 := O[25].14; //spare
   CB_1CS:1:O.15 := O[25].15; //spare
   
   // CROSSBREAK ZONE 2
   CB_2CS:1:O.0 := O[27].0; //CRSSBRK ZONE 2 North Outside Lamp
   CB_2CS:1:O.1 := O[27].1; //CRSSBRK ZONE 2 North Inside Lamp
   CB_2CS:1:O.2 := O[27].2; //CRSSBRK ZONE 2 South Outside Lamp (Bad Output)
   CB_2CS:1:O.3 := O[27].3; //CRSSBRK ZONE 2 South Inside Lamp
   CB_2CS:1:O.4 := O[27].4; //CRSSBRK ZONE 2 Crossbreak In progress Lamp
   CB_2CS:1:O.5 := O[27].5; //CRSSBRK ZONE 1 Crossbreak horn Located on wall At lehr Exit
   CB_2CS:1:O.6 := O[27].6; //CRSSBRK ZONE 1 Alarm rotating Beacon Located on lehr Exit
   CB_2CS:1:O.7 := O[27].7; //Crusher #1 Is Lowered (This Output is Read by HE for Pan-alarm Display)
   CB_2CS:1:O.8 := O[27].8; //CRSSBRK ZONE 2 South Outside Lamp (New Output)
   CB_2CS:1:O.9 := O[27].9; //spare
   CB_2CS:1:O.10 := O[27].10; //spare
   CB_2CS:1:O.11 := O[27].11; //spare
   CB_2CS:1:O.12 := O[27].12; //spare
   CB_2CS:1:O.13 := O[27].13; //spare
   CB_2CS:1:O.14 := O[27].14; //spare
   CB_2CS:1:O.15 := O[27].15; //spare
   
   // CROSSBREAK ZONE 3
   CB_3CS:1:O.0 := O[29].0; //CRSSBRK ZONE 3 North Outside Lamp
   CB_3CS:1:O.1 := O[29].1; //CRSSBRK ZONE 3 North Inside Lamp
   CB_3CS:1:O.2 := O[29].2; //CRSSBRK ZONE 3 South Outside Lamp (Bad Output)
   CB_3CS:1:O.3 := O[29].3; //CRSSBRK ZONE 3 South Inside Lamp
   CB_3CS:1:O.4 := O[29].4; //CRSSBRK ZONE 3 Crossbreak In progress Lamp
   CB_3CS:1:O.5 := O[29].5; //spare
   CB_3CS:1:O.6 := O[29].6; //spare
   CB_3CS:1:O.7 := O[29].7; //spare
   CB_3CS:1:O.8 := O[29].8; //spare
   CB_3CS:1:O.9 := O[29].9; //spare
   CB_3CS:1:O.10 := O[29].10; //spare
   CB_3CS:1:O.11 := O[29].11; //spare
   CB_3CS:1:O.12 := O[29].12; //spare
   CB_3CS:1:O.13 := O[29].13; //spare
   CB_3CS:1:O.14 := O[29].14; //spare
   CB_3CS:1:O.15 := O[29].15; //spare
   
   // CROSSBREAK ZONE 4 (IMAGE AUTO)
   CB_4CS:1:O.0 := O[31].0; //CRSSBRK ZONE 4 North Outside Lamp
   CB_4CS:1:O.1 := O[31].1; //CRSSBRK ZONE 4 North Inside Lamp
   CB_4CS:1:O.2 := O[31].2; //CRSSBRK ZONE 4 South Outside Lamp (Bad Output)
   CB_4CS:1:O.3 := O[31].3; //CRSSBRK ZONE 4 South Inside Lamp
   CB_4CS:1:O.4 := O[31].4; //CRSSBRK ZONE 4 Crossbreak In progress Lamp
   CB_4CS:1:O.5 := O[31].5; //spare
   CB_4CS:1:O.6 := O[31].6; //IMAGE AUTO Retro cover Manual  mode Lamp
   CB_4CS:1:O.7 := O[31].7; //IMAGE AUTO Retro cover Closed Alarm Horn
   CB_4CS:1:O.8 := O[31].8; //IMAGE AUTO Retro cover Alarm Beacon
   CB_4CS:1:O.9 := O[31].9; //IMAGE AUTO Open Graticule Solenoid (Raise)
   CB_4CS:1:O.10 := O[31].10; //IMAGE AUTO Retro Cover Open solenoid Valve
   CB_4CS:1:O.11 := O[31].11; //spare
   CB_4CS:1:O.12 := O[31].12; //spare
   CB_4CS:1:O.13 := O[31].13; //spare
   CB_4CS:1:O.14 := O[31].14; //spare
   CB_4CS:1:O.15 := O[31].15; //spare
   
   // CROSSBREAK ZONE 5 (APC)
   CB_5CS:1:O.0 := O[33].0; //CRSSBRK ZONE 5 North Outside Lamp
   CB_5CS:1:O.1 := O[33].1; //CRSSBRK ZONE 5 North Inside Lamp
   CB_5CS:1:O.2 := O[33].2; //CRSSBRK ZONE 5 South Outside Lamp (Bad Output)
   CB_5CS:1:O.3 := O[33].3; //CRSSBRK ZONE 5 South Inside Lamp
   CB_5CS:1:O.4 := O[33].4; //CRSSBRK ZONE 5 Crossbreak In progress Lamp
   CB_5CS:1:O.5 := O[33].5; //APC Enable Relay
   CB_5CS:1:O.6 := O[33].6; //APC Cut Off relay New Apc Sprayer
   CB_5CS:1:O.7 := O[33].7; //APC #2 Blow off Excess APC During Crossbreak
   CB_5CS:1:O.8 := O[33].8; //APC #2 Lower Roll (On Glass)
   CB_5CS:1:O.9 := O[33].9; //APC #1 Blow off Excess APC During Crossbreak changed 22Mar2019TC
   CB_5CS:1:O.10 := O[33].10; //APC #1 Lower Roll (On Glass) new22MarTC
   CB_5CS:1:O.11 := O[33].11; //APC APC Roll SS1 changed 22Mar2019TC
   CB_5CS:1:O.12 := O[33].12; //spare
   CB_5CS:1:O.13 := O[33].13; //spare
   CB_5CS:1:O.14 := O[33].14; //spare
   CB_5CS:1:O.15 := O[33].15; //spare
   
   // MANUAL INSPECTION
   MI_6CS:1:O.0 := O[35].0; //MANUAL INSPCTN North Outside Reject Flaw Red Lamp
   MI_6CS:1:O.1 := O[35].1; //MANUAL INSPCTN North Outside Q.A. Flaw Yellow Lamp
   MI_6CS:1:O.2 := O[35].2; //MANUAL INSPCTN North Inside Reject Flaw Red Lamp
   MI_6CS:1:O.3 := O[35].3; //MANUAL INSPCTN North Inside Q.A. Flaw Yellow Lamp
   MI_6CS:1:O.4 := O[35].4; //MANUAL INSPCTN * Center Reject Flaw Red Lamp
   MI_6CS:1:O.5 := O[35].5; //MANUAL INSPCTN * Center Q.A. Flaw Yellow Lamp
   MI_6CS:1:O.6 := O[35].6; //MANUAL INSPCTN South Inside Reject Flaw Red Lamp
   MI_6CS:1:O.7 := O[35].7; //MANUAL INSPCTN South Inside Q.A. Flaw Yellow Lamp
   MI_6CS:1:O.8 := O[35].8; //MANUAL INSPCTN South Outside Reject Flaw Red Lamp
   MI_6CS:1:O.9 := O[35].9; //MANUAL INSPCTN South Outside Q.A. Flaw Yellow Lamp
   MI_6CS:1:O.10 := O[35].10; //MANUAL INSPCTN Cross-break Signal to STP
   MI_6CS:1:O.11 := O[35].11; //spare
   MI_6CS:1:O.12 := O[35].12; //spare
   MI_6CS:1:O.13 := O[35].13; //MANUAL INSPCTN * * Function Lamp Clear
   MI_6CS:1:O.14 := O[35].14; //MANUAL INSPCTN * * Function Lamp Blue
   MI_6CS:1:O.15 := O[35].15; //MANUAL INSPCTN Quality Defect Inhibit Function Lamp Red
   
   //Cabinet
   A152AP1:15:O.Pt15.Data := TMP_xSimulationMode; //PLC ANOMALY
   A152AP1:17:O.Pt00.Data := O[35].15; //MANUAL INSPECTION
   
   //VMCC W1 (WASHER)
   
   
   
   //PANEL W2 (WASHER)
   PANEL_W2:3:O.0 := O[59].0; //PANEL W2 BRUSH #1 Manual mode Lamp
   PANEL_W2:3:O.1 := O[59].1; //SPARE
   PANEL_W2:3:O.2 := O[59].2; //PANEL W2 SPONGE UNIT Manual mode Lamp
   PANEL_W2:3:O.3 := O[59].3; //PANEL W2 AIR KNIVES Manual mode Lamp
   PANEL_W2:3:O.4 := O[59].4; //PANEL W2 WATER SPRAYERS Manual mode Lamp
   PANEL_W2:3:O.5 := O[59].5; //SPARE
   PANEL_W2:3:O.6 := O[59].6; //PANEL W2 AIR KNIFE SS LIGHT ON PANEL #W2
   PANEL_W2:3:O.7 := O[59].7; //PANEL W2 AIR KNIFE RELAY AKBR-ON
   PANEL_W2:3:O.8 := O[59].8; //SPARE
   PANEL_W2:3:O.9 := O[59].9; //SPARE
   PANEL_W2:3:O.10 := O[59].10; //SPARE
   PANEL_W2:3:O.11 := O[59].11; //SPARE
   PANEL_W2:3:O.12 := O[59].12; //SPARE
   PANEL_W2:3:O.13 := O[59].13; //SPARE
   PANEL_W2:3:O.14 := O[59].14; //SPARE
   PANEL_W2:3:O.15 := O[59].15; //SPARE
   
   //PANEL W3 (WASHER)
   PANEL_W3:3:O.0 := O[63].0; //PANEL W3 BRUSH #1 Manual mode Lamp
   PANEL_W3:3:O.1 := O[63].1; //SPARE
   PANEL_W3:3:O.2 := O[63].2; //PANEL W3 SPONGE UNIT Manual mode Lamp
   PANEL_W3:3:O.3 := O[63].3; //PANEL W3 AIR KNIVES Manual mode Lamp
   PANEL_W3:3:O.4 := O[63].4; //PANEL W3 WATER SPRAYERS Manual mode Lamp
   PANEL_W3:3:O.5 := O[63].5; //SPARE
   PANEL_W3:3:O.6 := O[63].6; //PANEL W3 AIR KNIFE SS LIGHT ON PANEL #W3
   PANEL_W3:3:O.7 := O[63].7; //SPARE
   PANEL_W3:3:O.8 := O[63].8; //SPARE
   PANEL_W3:3:O.9 := O[63].9; //SPARE
   PANEL_W3:3:O.10 := O[63].10; //SPARE
   PANEL_W3:3:O.11 := O[63].11; //SPARE
   PANEL_W3:3:O.12 := O[63].12; //SPARE
   PANEL_W3:3:O.13 := O[63].13; //SPARE
   PANEL_W3:3:O.14 := O[63].14; //SPARE
   PANEL_W3:3:O.15 := O[63].15; //SPARE
   
   
   //PRODUCED
   
   To_Cullet[0] := O[112];
   To_Cullet[1] := O[113];
   To_Cullet[2] := O[114];
   To_Cullet[3] := O[115];
   To_Cullet[4] := O[116];
   To_Cullet[5] := O[117];
   To_Cullet[6] := O[118];
   To_Cullet[7] := O[119];
   
   /*
   
   ProducedToCullet.MBtoCULLET_1 := O[112];
   ProducedToCullet.MBtoCULLET_2 := O[113];
   ProducedToCullet.MBtoCULLET_3 := O[114];
   ProducedToCullet.MBtoCULLET_4 := O[115];
   ProducedToCullet.MBtoCULLET_5 := O[116];
   ProducedToCullet.MBtoCULLET_6 := O[117];
   ProducedToCullet.MBtoCULLET_7 := O[118];
   ProducedToCullet.MBtoCULLET_8 := O[119];
   
   */
   
   ProducedToMCC1300.iMBtoM2_1 := O[120];
   ProducedToMCC1300.iMBtoM2_2 := O[121];
   ProducedToMCC1300.iMBtoM2_3 := O[122];
   ProducedToMCC1300.iMBtoM2_4 := O[123];
   ProducedToMCC1300.iMBtoM2_5 := O[124];
   ProducedToMCC1300.iMBtoM2_6 := O[125];
   ProducedToMCC1300.iMBtoM2_7 := O[126];
   ProducedToMCC1300.iMBtoM2_8 := O[127];
   
   
   //DRIVE
   
   
END_ROUTINE

ROUTINE _9_SPEED_CON   (* ladder *)